// TIA Portal project "XSFW_TIA60401_A5" (V13) (continued)
   "ArrMC005" AT %T79 : Timer;   // Timer arranque MC005
   "MC004_TTB" AT %E6.3 : Bool;   // M COMPRESOR ALTA ABC4-TERMOSTATO AGUA / Compresor ABC4 Alta Temperatura de agua
   "MC005" AT %A1.2 : Bool;   // M COMPRESOR ALTA ABC5-CONTACTOR / Compresor ABC5-. Marcha-(200 Kw)
   "MC005-CO" AT %E3.5 : Bool;   // M COMPRESOR ALTA ABC5-CONFIRMACIÓN DE MARCHA / Compresor ABC5-Confirmacion Marcha-(200 Kw)
   "MC005-TO" AT %E3.6 : Bool;   // M COMPRESOR ALTA ABC5-TÉRMICO / Compresor ABC5-Falla Termico--(200 Kw)
   "MC005_EV" AT %A2.4 : Bool;   // M COMPRESOR ALTA ABC5-ELECTROVÁLVULA / Electrovalvula libera carga MC005 (ABC5)
   "MC005_MANT" AT %A3.1 : Bool;   // M COMPRESOR ALTA ABC5-SEÑAL MODO MANTENIMIENTO / Compresor MC005 Salida Mantenimiento
   "MC005_PTA" AT %E6.4 : Bool;   // M COMPRESOR ALTA ABC5-PRESOSTATO ACEITE / Compresor ABC5 Baja Presion de Aceite
   "MC005_PTB" AT %E6.5 : Bool;   // M COMPRESOR ALTA ABC5-PRESOSTATO AGUA / Compresor ABC5 Baja Presion de Agua
   "MC005_TTA" AT %E6.6 : Bool;   // M COMPRESOR ALTA ABC5-TERMOSTATO AIRE / Compresor ABC5 Alta Temperatura de Aire
   "MC005_TTB" AT %E6.7 : Bool;   // M COMPRESOR ALTA ABC5-TERMOSTATO AGUA / Compresor ABC5 Alta Temperatura de agua
   "MC060-CO" AT %E10.0 : Bool;   // M COMPR BAJA SULLAIR 2-CONFIRMACIÓN DE MARCHA / Compresor Baja XXX - Conf.Marcha
   "MC060-TO" AT %E10.1 : Bool;   // M COMPR BAJA SULLAIR 2-TÉRMICO / Compresor Baja XXX - Falla de termico
   "MC060-VS1" AT %E10.2 : Bool;   // M COMPR BAJA SULLAIR 2-PULSADOR PARADA / Compresor Baja XXX - Falla de seguridades
   "MC060_MANT" AT %A5.4 : Bool;   // M COMPR BAJA SULLAIR 2-SEÑAL MODO MANTENIMIENTO / compresor XXX salida de mantenimiento
   "MC060_MARCHA" AT %A5.5 : Bool;   // M COMPR BAJA SULLAIR 2-CONTACTOR / compresor XXX salida de marcha
   "MC061-CO" AT %E11.4 : Bool;   // M COMPR BAJA SULLAIR 1-CONFIRMACIÓN DE MARCHA / Compresor Baja SULL 1 - Conf.Marcha
   "MC003_EV" AT %A2.2 : Bool;   // M COMPRESOR ALTA BELLIS-ELECTROVÁLVULA 1 / Electrovalvula libera carga MC003 (Bellis)
   "Encendido" AT %M301.1 : Bool;   // Encendido de PLC
   "MT009-TO" AT %E66.5 : Bool;   // B INT L3 Y L5-TÉRMICO / Bomba Principal Chiller Envasado - Falla de Térmico
   "MT010-CO" AT %E66.6 : Bool;   // B INT L1 Y MANOMEC-CONFIRMACIÓN DE MARCHA / Bomba Auxilliar Chiller Envasado - Confirmación de Marcha
   "MT010-Marcha" AT %A66.3 : Bool;   // B INT L1 Y MANOMEC-CONTACTOR / Accionamiento Bomba Intercambiador LINEA 1 Y MANOMEC
   "MT010-TO" AT %E66.7 : Bool;   // B INT L1 Y MANOMEC-TÉRMICO / Bomba Auxiliar Chiller Envasado - Falla de Térmico
   "MV030" AT %A0.2 : Bool;   // M VENTILADOR 2-CONTACTOR / VENTILADOR TORRE 1 -. marcha-
   "MV030-CO" AT %E0.4 : Bool;   // M VENTILADOR 2-CONFIRMACIÓN DE MARCHA / VENTILADOR TORRE 1 -confirmacion marcha-
   "MV030-TO" AT %E0.5 : Bool;   // M VENTILADOR 2-TÉRMICO / VENTILADOR TORRE 1 -falla termico-
   "MV030_PA" AT %E8.5 : Bool;   // M VENTILADOR 2-PULSADOR MARCHA / Ventilador 1 Torre Cavalleto Pulsador Arranque
   "MV030_PP" AT %E8.6 : Bool;   // M VENTILADOR 2-PULSADOR PARADA / Ventilador 1 Torre Cavalleto Pulsador Parada
   "MV031" AT %A0.3 : Bool;   // M VENTILADOR 1-CONTACTOR / VENTILADOR TORRE 2 -. marcha-
   "MV031-CO" AT %E0.6 : Bool;   // M VENTILADOR 1-CONFIRMACIÓN DE MARCHA / VENTILADOR TORRE 2 -confirmacion marcha-
   "MV031-TO" AT %E0.7 : Bool;   // M VENTILADOR 1-TÉRMICO / VENTILADOR TORRE 2 -falla termico-
   "MV031_PA" AT %E8.7 : Bool;   // M VENTILADOR 1-PULSADOR MARCHA / Ventilador 2 Torre Cavalleto Pulsaor Arranque
   "MV031_PP" AT %E9.0 : Bool;   // M VENTILADOR 1-PULSADOR PARADA / Ventilador 2 Torre Cavalleto Pulsaor Parada
   "iGMBooster2" AT %E9.7 : Bool;   // M BOOSTER 2-GUARDAMOTOR / Guardamotor Booster 2
   "Hab-CHILL1" AT %A69.4 : Bool;   // CHILLER 1-SEÑAL A CHILLER / Deshabilitación Chiller Soplado GRANDE
   "Hab-CHILL2" AT %A69.5 : Bool;   // CHILLER 2-SEÑAL A CHILLER / Deshabilitación Chiller Soplado CHICO
   "Hab-CHILL3" AT %A69.6 : Bool;   // CHILLER 3-SEÑAL A CHILLER / Deshabilitación Chiller Envasado GRANDE
   "Hab-CHILL4" AT %A69.7 : Bool;   // CHILLER 4-SEÑAL A CHILLER / Deshabilitación Chiller Envasado CHICO
   "ILUMINACION" AT %A0.5 : Bool;   // ILUMINACION-CONTACTOR / ILUMINACION
   "MC003_ConfPurga" AT %E1.2 : Bool;   // Bellis - Confirmación de electroválvula de purga. / Iluminacion-confirmacion marcha-
   "MC004_ConfPurga" AT %E1.3 : Bool;   // ABC4 - Confirmación de electroválvula de purga. / Iluminacion Termico
   "IndicadorChillers" AT %M310.0 : Bool;   // Indicador Aviso en chillers
   "TsinReq1" AT %T52 : Timer;   // Timeout estando en estado sin requerimiento 1
   "TsinReq2" AT %T40 : Timer;   // Timeout estando en estado sin requerimiento 2
   "TsinReq3" AT %T41 : Timer;   // Timeout estando en estado sin requerimiento 3
   "TsinReq4" AT %T42 : Timer;   // Timeout estando en estado sin requerimiento 4
   "TsinReq5" AT %T43 : Timer;   // Timeout estando en estado sin requerimiento 5
   "UNO" AT %M0.1 : Bool;
   "V001-CO" AT %E76.5 : Bool;   // VENT 1 TORR ENF CHILLERS-CONFIRMACIÓN DE MARCHA / Ventilador 1 Torres Enfriamiento - Confirmación de Marcha
   "V001-Marcha" AT %A67.6 : Bool;   // VENT 1 TORR ENF CHILLERS-CONTACTOR / Accionamiento Ventilador 1 Torres Enfriamiento
   "V001-TO" AT %E76.6 : Bool;   // VENT 1 TORR ENF CHILLERS-TÉRMICO / Ventilador 1 Torres Enfriamiento - Falla de Térmico
   "V002-CO" AT %E76.7 : Bool;   // VENT 2 TORR ENF CHILLERS-CONFIRMACIÓN DE MARCHA / Ventilador 2 Torres Enfriamiento - Confirmación de Marcha
   "V002-Marcha" AT %A67.7 : Bool;   // VENT 2 TORR ENF CHILLERS-CONTACTOR / Accionamiento Ventilador 2 Torres Enfriamiento
   "V002-TO" AT %E77.0 : Bool;   // VENT 2 TORR ENF CHILLERS-TÉRMICO / Ventilador 2 Torres Enfriamiento - Falla de Térmico
   "V003-CO" AT %E77.1 : Bool;   // VENT 3 TORR ENF CHILLERS-CONFIRMACIÓN DE MARCHA / Ventilador 3 Torres Enfriamiento - Confirmación de Marcha
   "V003-Marcha" AT %A68.0 : Bool;   // VENT 3 TORR ENF CHILLERS-CONTACTOR / Accionamiento Ventilador 3 Torres Enfriamiento
   "V003-TO" AT %E77.2 : Bool;   // VENT 3 TORR ENF CHILLERS-TÉRMICO / Ventilador 3 Torres Enfriamiento - Falla de Térmico
   "FlancoNSop1" AT %M326.1 : Bool;
   "FlancoNSop2" AT %M326.2 : Bool;
   "FlancoNSop3" AT %M326.3 : Bool;
   "FlancoNoFaGen" AT %M325.2 : Bool;
   "FlancoNoFal1" AT %M324.5 : Bool;
   "MC003_EV2" AT %A3.2 : Bool;   // M COMPRESOR ALTA BELLIS-ELECTROVÁLVULA 2 / Electrovalvula media carga Bellis
   "MC003_FTA" AT %E7.4 : Bool;   // M COMPRESOR ALTA BELLIS-FUJOSTATO / Compresor Bellis & MHW28 Falla de Flujostato
   "MC003_MANT" AT %A2.7 : Bool;   // M COMPRESOR ALTA BELLIS-SEÑAL MODO MANTENIMIENTO / Compresor MC003 Salida Mantenimiento
   "MC003_PTA" AT %E7.0 : Bool;   // M COMPRESOR ALTA BELLIS-PRESOSTATO ACEITE / Compresor Bellis & MHW28 Baja Presion Aceite
   "MC003_PTB" AT %E7.1 : Bool;   // M COMPRESOR ALTA BELLIS-PRESOSTATO AGUA / Compresor Bellis & MHW28 Baja Presion de Agua
   "MC003_TTA" AT %E7.2 : Bool;   // M COMPRESOR ALTA BELLIS-TERMOSTATO AIRE / Compresor Bellis & MHW28 Alta temperatura de Aire
   "MC003_TTB" AT %E7.3 : Bool;   // M COMPRESOR ALTA BELLIS-TERMOSTATO AGUA / Compresor Bellis & MHW28 Alta temperatura de Agua
   "MC004" AT %A1.1 : Bool;   // M COMPRESOR ALTA ABC4-CONTACTOR / Compresor ABC4-. Marcha-
   "MC004-CO" AT %E3.3 : Bool;   // M COMPRESOR ALTA ABC4-CONFIRMACIÓN DE MARCHA / Compresor ABC4-Confirmacion Marcha-
   "MC004-TO" AT %E3.4 : Bool;   // M COMPRESOR ALTA ABC4-TÉRMICO / Compresor ABC4-Falla Termico-
   "MC004_EV" AT %A2.3 : Bool;   // M COMPRESOR ALTA ABC4-ELECTROVÁLVULA / Electrovalvula libera carga MC004 (ABC4)
   "MC004_MANT" AT %A3.0 : Bool;   // M COMPRESOR ALTA ABC4-SEÑAL MODO MANTENIMIENTO / Compresor MC004 Salida Mantenimiento
   "MC004_PTA" AT %E6.0 : Bool;   // M COMPRESOR ALTA ABC4-PRESOSTATO ACEITE / Compresor ABC4 Baja Presion de Aceite
   "MC004_PTB" AT %E6.1 : Bool;   // M COMPRESOR ALTA ABC4-PRESOSTATO AGUA / Compresor ABC4 Baja Presion de Agua
   "MC004_TTA" AT %E6.2 : Bool;   // M COMPRESOR ALTA ABC4-TERMOSTATO AIRE / Compresor ABC4 Alta Temperatura de Aire
   "MC001_PTA" AT %E5.0 : Bool;   // M COMPRESOR ALTA ABC2-PRESOSTATO ACEITE / Compresor ABC2 Baja Presion de Aceite
   "MC001_PTB" AT %E5.1 : Bool;   // M COMPRESOR ALTA ABC2-PRESOSTATO AGUA / Compresor ABC2 Baja Presion de Agua
   "MC001_TTA" AT %E5.2 : Bool;   // M COMPRESOR ALTA ABC2-TERMOSTATO AIRE / Compresor ABC2 Alta Temperatura de Aire
   "MC001_TTB" AT %E5.3 : Bool;   // M COMPRESOR ALTA ABC2-TERMOSTATO AGUA / Compresor ABC2 Alta Temperatura de agua
   "MC002" AT %A0.7 : Bool;   // M COMPRESOR ALTA ABC3-CONTACTOR / Compresor ABC3-. Marcha-
   "MC002-CO" AT %E2.7 : Bool;   // M COMPRESOR ALTA ABC3-CONFIRMACIÓN DE MARCHA / Compresor ABC3-Confirmacion Marcha-
   "MC002-TO" AT %E3.0 : Bool;   // M COMPRESOR ALTA ABC3-TÉRMICO / Compresor ABC3-Falla Termico-
   "MC002_EV" AT %A2.1 : Bool;   // M COMPRESOR ALTA ABC3-ELECTROVÁLVULA / Electrovalvula libera carga MC002 (ABC3)
   "MC002_MANT" AT %A2.6 : Bool;   // M COMPRESOR ALTA ABC3-SEÑAL MODO MANTENIMIENTO / Compresor MC002 Salida Mantenimiento
   "MC002_PTA" AT %E5.4 : Bool;   // M COMPRESOR ALTA ABC3-PRESOSTATO ACEITE / Compresor ABC3 Baja Presion de Aceite
   "MC002_PTB" AT %E5.5 : Bool;   // M COMPRESOR ALTA ABC3-PRESOSTATO AGUA / Compresor ABC3 Baja Presion de Agua
   "MC002_TTA" AT %E5.6 : Bool;   // M COMPRESOR ALTA ABC3-TERMOSTATO AIRE / Compresor ABC3 Alta Temperatura de Aire
   "MC002_TTB" AT %E5.7 : Bool;   // M COMPRESOR ALTA ABC3-TERMOSTATO AGUA / Compresor ABC3 Alta Temperatura de agua
   "MC003" AT %A1.0 : Bool;   // M COMPRESOR ALTA BELLIS-CONTACTOR / Compresor B&MWH28-. Marcha-
   "MC003-CO" AT %E3.1 : Bool;   // M COMPRESOR ALTA BELLIS-CONFIRMACIÓN DE MARCHA / Compresor B&MWH28-Confirmacion Marcha-
   "MC003-TO" AT %E3.2 : Bool;   // M COMPRESOR ALTA BELLIS-TÉRMICO / Compresor B&MWH28-Falla Termico-
   "BoostPlsManual" AT %M10.6 : Bool;   // Booster Pulsa Manual desde HMI
   "BoostPlsAutoma" AT %M10.7 : Bool;   // Booster Pulsa Automático desde HMI
   "ErrPMQG" AT %M321.2 : Bool;   // Error Prioritarias General
   "PRESOSTATO-TORRES" AT %E76.4 : Bool;   // CHILLER (TODOS)-PRESOSTATO / Presostato Agua Torres de Enfriamiento
   "PT2_AIRE" AT %E4.7 : Bool;   // - / PRESOSTATO ALTA PRESION DE AIRE EN COLECTOR 40Kg
   "Parada-MC061" AT %A6.1 : Bool;   // M COMPR BAJA SULLAIR 1-ORDEN PARADA / Parada MC061
   "MC006_ConfPurga" AT %E11.7 : Bool;   // ABC1 - Confirmación de electroválvula de purga.
   "MP014-TO" AT %E0.1 : Bool;   // BOMBA 1-TÉRMICO / BOMBA 1TORRE ENF.-TERMICO
   "MP015" AT %A0.1 : Bool;   // BOMBA 2-CONTACTOR / BOMBA 2 TORRE -. marcha-
   "MP015-CO" AT %E0.2 : Bool;   // BOMBA 2-CONFIRMACIÓN DE MARCHA / BOMBA 2 TORRE ENF.-CONFIRMACION
   "MP015-TO" AT %E0.3 : Bool;   // BOMBA 2-TÉRMICO / BOMBA 2 TORRE ENF.-TERMICO
   "MP018-CO" AT %E68.0 : Bool;   // BOMBA 1-CONFIRMACIÓN DE MARCHA / Bomba 1 Torres Enfriamiento - Confirmación de Marcha
   "MP018-Marcha" AT %A67.0 : Bool;   // BOMBA 1-CONTACTOR / Accionamiento Bomba 1 Torres Enfriamiento
   "MP018-TO" AT %E68.1 : Bool;   // BOMBA 1-TÉRMICO / Bomba 1 Torres Enfriamiento - Falla de Térmico
   "MP018_PA" AT %E8.1 : Bool;   // BOMBA 1-PULSADOR MARCHA / Bomba 1 Torre Cavalleto Pulsador Arranque
   "MP018_PP" AT %E8.2 : Bool;   // BOMBA 1-PULSADOR PARADA / Bomba 1 Torre Cavalleto Pulsador Parada
   "MC001_ConfPurga" AT %E1.0 : Bool;   // ABC2 - Confirmación de electroválvula de purga. / Bomba de pozo -confirmacion marcha-
   "CERO" AT %M0.0 : Bool;
   "CHILL1-AL1" AT %E68.4 : Bool;   // CHILLER SOPLADO-ALARMA 1 / Chiller Soplado GRANDE - Alarma 1
   "CHILL1-AL2" AT %E68.5 : Bool;   // CHILLER SOPLADO-ALARMA 2 / Chiller Soplado GRANDE - Alarma 2
   "CHILL1-MAX" AT %E68.7 : Bool;   // CHILLER SOPLADO-MAXIMA CAPACIDAD / Chiller Soplado GRANDE - Máxima Capacidad
   "CHILL1-RUN" AT %E68.6 : Bool;   // CHILLER SOPLADO- / Chiller Soplado GRANDE - En modo RUN
   "CHILL2-" AT %E69.0 : Bool;   // CHILLER SOPLADO CHICO- / Chiller Soplado CHICO - Contactor 1
   "CHILL2-b" AT %E69.1 : Bool;   // CHILLER SOPLADO CHICO- / Chiller Soplado CHICO - Contactor 2
   "CHILL2-c" AT %E69.2 : Bool;   // CHILLER SOPLADO CHICO-FALLA / Chiller Soplado CHICO - Termico Contactor 1
   "CHILL2-d" AT %E69.3 : Bool;   // CHILLER SOPLADO CHICO-FALLA / Chiller Soplado CHICO - Termico Contactor 2
   "CHILL3-AL1" AT %E69.4 : Bool;   // CHILLER ENVASADO GRAND-ALARMA 1 / Chiller Envasado GRANDE - Alarma 1
   "MC064-VS1" AT %E11.3 : Bool;   // M COMPR BAJA ATLAS 2-PULSADOR PARADA / Compresor Baja ATLAS 2 - Falla de seguridades
   "MC064_MANT" AT %A5.2 : Bool;   // M COMPR BAJA ATLAS 2-SEÑAL MODO MANTENIMIENTO / compresor ATLAS 2 salida de mantenimiento
   "MC064_MARCHA" AT %A5.3 : Bool;   // M COMPR BAJA ATLAS 2-CONTACTOR / compresor ATLAS 2 salida de marcha
   "MP010-CO" AT %E67.0 : Bool;   // B PRINC CH. SOPLADO-CONFIRMACIÓN DE MARCHA / Bomba Intercambiador LINEA 1 - Confirmación de Marcha
   "MP010-Marcha" AT %A66.4 : Bool;   // B PRINC CH. SOPLADO-CONTACTOR / Accionamiento Bomba Principal Chiller Soplado
   "MP010-TO" AT %E67.1 : Bool;   // B PRINC CH. SOPLADO-TÉRMICO / Bomba Intercambiador LINEA 1 - Falla de Térmico
   "MC006" AT %Q6.2 : Bool;   // M COMPRESOR ALTA ABC1-CONTACTOR
   "MC006_EV" AT %Q6.3 : Bool;   // M COMPRESOR ALTA ABC1-ELECTROVÁLVULA
   "MC006_MANT" AT %Q6.4 : Bool;   // M COMPRESOR ALTA ABC1-SEÑAL MODO MANTENIMIENTO
   "TsinReq6" AT %T59 : Timer;
   "TV6" AT %T69 : Timer;
   "flReqMch6" AT %M0.5 : Bool;
   "ErrPMQ6" AT %M1.5 : Bool;
   "ErrCMQ6" AT %M1.6 : Bool;
   "RetVLV6" AT %T85 : Timer;
   "TRetVCmp6" AT %T86 : Timer;
   "ArrMC006" AT %T88 : Timer;
   "FlaAux6" AT %M301.2 : Bool;
   "FlancoINC6" AT %M326.7 : Bool;
   "FlancoDEC6" AT %M327.0 : Bool;
   "FlancoMan6" AT %M327.1 : Bool;
   "FlancoManP6" AT %M327.2 : Bool;
   "FlancoAuto6" AT %M327.3 : Bool;
   "FlancoNoFal6" AT %M327.4 : Bool;
   "FlancoTSinReq6" AT %M327.5 : Bool;
   "AuxTempMS050" AT %MW340 : Int;
   "AuxTempMS051" AT %MW342 : Int;
   "AuxTempMS052" AT %MW344 : Int;
   "AuxTempMS053" AT %MW346 : Int;
   "AuxTempMS054" AT %MW348 : Int;
   "AuxTempMS055" AT %MW350 : Int;
   "AuxTempMS056" AT %MW352 : Int;
   "AuxTempMC060" AT %MW354 : Int;
   "AuxTempMC061" AT %MW356 : Int;
   "AuxTempMC062" AT %MW358 : Int;
   "AuxTempMC063" AT %MW360 : Int;
   "AuxTempMC064" AT %MW362 : Int;
   "AuxTempMC065" AT %MW364 : Int;
   "ProxMantBoost1" AT %MD16 : DInt;
   "LimiteMantBoost1" AT %M1.7 : Bool;
   "ProxMantBoost2" AT %MD26 : DInt;
   "LimiteMantBoost2" AT %M2.3 : Bool;
END_VAR

DATA_BLOCK "DB_Fecha"   // DB1
{ S7_Optimized_Access := 'FALSE' }
VERSION : 0.1
   VAR
      STAT0 : Date_And_Time;
      STAT1 : Int;
      STAT2 : Int;
      STAT3 : Int;
      STAT4 : Int;
      STAT5 : Int;
      STAT6 : Int;
      STAT7 : Int;
      STAT8 : Int;
      STAT9 : Int;
      STAT10 : Int;
      STAT11 : Word;
      STAT12 : Word;
      STAT13 : Word;
      STAT14 : Word;
      STAT15 : Word;
      STAT16 : Word;
   END_VAR
BEGIN
END_DATA_BLOCK

DATA_BLOCK "Enclavamientos"   // DB28
{ S7_Optimized_Access := 'FALSE' }
VERSION : 0.1
   VAR
      En1 : Bool;
      En2 : Bool;
      En3 : Bool;
      En4 : Bool;
      En5 : Bool;
      En6 : Bool;
      En7 : Bool;
      En8 : Bool;
      En9 : Bool;
      En10 : Bool;
      En11 : Bool;
      En12 : Bool;
      En13 : Bool;
      En14 : Bool;
      En15 : Bool;
      En16 : Bool;
      En17 : Bool;
      En18 : Bool;
      En19 : Bool;
      En20 : Bool;
      En21 : Bool;
      En22 : Bool;
      En23 : Bool;
      En24 : Bool;
      En25 : Bool;
      En26 : Bool;
      En27 : Bool;
      En28 : Bool;
      En29 : Bool;
      En30 : Bool;
      En31 : Bool;
      En32 : Bool;
      En33 : Bool;
      En34 : Bool;
      En35 : Bool;
      En36 : Bool;
      En37 : Bool;
      En38 : Bool;
      En39 : Bool;
      En40 : Bool;
      En41 : Bool;
      En42 : Bool;
      En43 : Bool;
      En44 : Bool;
      En45 : Bool;
      En46 : Bool;
      En47 : Bool;
      En48 : Bool;
      En49 : Bool;
      En50 : Bool;
      En51 : Bool;
      En52 : Bool;
      En53 : Bool;
      En54 : Bool;
      En55 : Bool;
      En56 : Bool;
      En57 : Bool;
      En58 : Bool;
      En59 : Bool;
      En60 : Bool;
      En61 : Bool;
      En62 : Bool;
      En63 : Bool;
      En64 : Bool;
   END_VAR
BEGIN
END_DATA_BLOCK

// folder: Alarmas

DATA_BLOCK "DB_ALA_PRE"   // DB32
{ S7_Optimized_Access := 'FALSE' }
VERSION : 0.1
   VAR
      x : Bool;
      x1 : Bool;
      x2 : Bool;
      x3 : Bool;
      x4 : Bool;
      x5 : Bool;
      x6 : Bool;
      x7 : Bool;
      x8 : Bool;
      x9 : Bool;
      x10 : Bool;
      x11 : Bool;
      x12 : Bool;
      x13 : Bool;
      x14 : Bool;
      x15 : Bool;
      x16 : Bool;
      x17 : Bool;
      x18 : Bool;
      x19 : Bool;
      x20 : Bool;
      x21 : Bool;
      x22 : Bool;
      x23 : Bool;
      x24 : Bool;
      x25 : Bool;
      x26 : Bool;
      x27 : Bool;
      x28 : Bool;
      x29 : Bool;
      x30 : Bool;
      x31 : Bool;
      x32 : Bool;
      x33 : Bool;
      x34 : Bool;
      x35 : Bool;
      x36 : Bool;
      x37 : Bool;
      x38 : Bool;
      x39 : Bool;
      x40 : Bool;
      x41 : Bool;
      x42 : Bool;
      x43 : Bool;
      x44 : Bool;
      x45 : Bool;
      x46 : Bool;
      x47 : Bool;
      x48 : Bool;
      x49 : Bool;
      x50 : Bool;
      x51 : Bool;
      x52 : Bool;
      x53 : Bool;
      x54 : Bool;
      x55 : Bool;
      x56 : Bool;
      x57 : Bool;
      x58 : Bool;
      x59 : Bool;
      x60 : Bool;
      x61 : Bool;
      x62 : Bool;
      x63 : Bool;
      x64 : Bool;
      x65 : Bool;
      x66 : Bool;
      x67 : Bool;
      x68 : Bool;
      x69 : Bool;
      x70 : Bool;
      x71 : Bool;
      x72 : Bool;
      x73 : Bool;
      x74 : Bool;
      x75 : Bool;
      x76 : Bool;
      x77 : Bool;
      x78 : Bool;
      x79 : Bool;
      x80 : Bool;
      x81 : Bool;
      x82 : Bool;
      x83 : Bool;
      x84 : Bool;
      x85 : Bool;
      x86 : Bool;
      x87 : Bool;
      x88 : Bool;
      x89 : Bool;
      x90 : Bool;
      x91 : Bool;
      x92 : Bool;
      x93 : Bool;
      x94 : Bool;
      x95 : Bool;
      x96 : Bool;
      x97 : Bool;
      x98 : Bool;
      x99 : Bool;
      x100 : Bool;
      x101 : Bool;
      x102 : Bool;
      x103 : Bool;
      x104 : Bool;
      x105 : Bool;
      x106 : Bool;
      x107 : Bool;
      x108 : Bool;
      x109 : Bool;
      x110 : Bool;
      x111 : Bool;
      x112 : Bool;
      x113 : Bool;
      x114 : Bool;
      x115 : Bool;
      x116 : Bool;
      x117 : Bool;
      x118 : Bool;
      x119 : Bool;
      x120 : Bool;
      x121 : Bool;
      x122 : Bool;
      x123 : Bool;
      x124 : Bool;
      x125 : Bool;
      x126 : Bool;
      x127 : Bool;
      x128 : Bool;
      x129 : Bool;
      x130 : Bool;
      x131 : Bool;
      x132 : Bool;
      x133 : Bool;
      x134 : Bool;
      x135 : Bool;
      x136 : Bool;
      x137 : Bool;
      x138 : Bool;
      x139 : Bool;
      x140 : Bool;
      x141 : Bool;
      x142 : Bool;
      x143 : Bool;
      x144 : Bool;
      x145 : Bool;
      x146 : Bool;
      x147 : Bool;
      x148 : Bool;
      x149 : Bool;
      x150 : Bool;
      x151 : Bool;
      x152 : Bool;
      x153 : Bool;
      x154 : Bool;
      x155 : Bool;
      x156 : Bool;
      x157 : Bool;
      x158 : Bool;
      x159 : Bool;
      x160 : Bool;
      x161 : Bool;
      x162 : Bool;
      x163 : Bool;
      x164 : Bool;
      x165 : Bool;
      x166 : Bool;
      x167 : Bool;
      x168 : Bool;
      x169 : Bool;
      x170 : Bool;
      x171 : Bool;
      x172 : Bool;
      x173 : Bool;
      x174 : Bool;
      x175 : Bool;
      x176 : Bool;
      x177 : Bool;
      x178 : Bool;
      x179 : Bool;
      x180 : Bool;
      x181 : Bool;
      x182 : Bool;
      x183 : Bool;
      x184 : Bool;
      x185 : Bool;
      x186 : Bool;
      x187 : Bool;
      x188 : Bool;
      x189 : Bool;
      x190 : Bool;
      x191 : Bool;
      x192 : Bool;
      x193 : Bool;
      x194 : Bool;
      x195 : Bool;
      x196 : Bool;
      x197 : Bool;
      x198 : Bool;
      x199 : Bool;
   END_VAR
BEGIN
END_DATA_BLOCK

DATA_BLOCK "DB_ALA_REC"   // DB33
{ S7_Optimized_Access := 'FALSE' }
VERSION : 0.1
   VAR
      x : Bool;
      x1 : Bool;
      x2 : Bool;
      x3 : Bool;
      x4 : Bool;
      x5 : Bool;
      x6 : Bool;
      x7 : Bool;
      x8 : Bool;
      x9 : Bool;
      x10 : Bool;
      x11 : Bool;
      x12 : Bool;
      x13 : Bool;
      x14 : Bool;
      x15 : Bool;
      x16 : Bool;
      x17 : Bool;
      x18 : Bool;
      x19 : Bool;
      x20 : Bool;
      x21 : Bool;
      x22 : Bool;
      x23 : Bool;
      x24 : Bool;
      x25 : Bool;
      x26 : Bool;
      x27 : Bool;
      x28 : Bool;
      x29 : Bool;
      x30 : Bool;
      x31 : Bool;
      x32 : Bool;
      x33 : Bool;
      x34 : Bool;
      x35 : Bool;
      x36 : Bool;
      x37 : Bool;
      x38 : Bool;
      x39 : Bool;
      x40 : Bool;
      x41 : Bool;
      x42 : Bool;
      x43 : Bool;
      x44 : Bool;
      x45 : Bool;
      x46 : Bool;
      x47 : Bool;
      x48 : Bool;
      x49 : Bool;
      x50 : Bool;
      x51 : Bool;
      x52 : Bool;
      x53 : Bool;
      x54 : Bool;
      x55 : Bool;
      x56 : Bool;
      x57 : Bool;
      x58 : Bool;
      x59 : Bool;
      x60 : Bool;
      x61 : Bool;
      x62 : Bool;
      x63 : Bool;
      x64 : Bool;
      x65 : Bool;
      x66 : Bool;
      x67 : Bool;
      x68 : Bool;
      x69 : Bool;
      x70 : Bool;
      x71 : Bool;
      x72 : Bool;
      x73 : Bool;
      x74 : Bool;
      x75 : Bool;
      x76 : Bool;
      x77 : Bool;
      x78 : Bool;
      x79 : Bool;
      x80 : Bool;
      x81 : Bool;
      x82 : Bool;
      x83 : Bool;
      x84 : Bool;
      x85 : Bool;
      x86 : Bool;
      x87 : Bool;
      x88 : Bool;
      x89 : Bool;
      x90 : Bool;
      x91 : Bool;
      x92 : Bool;
      x93 : Bool;
      x94 : Bool;
      x95 : Bool;
      x96 : Bool;
      x97 : Bool;
      x98 : Bool;
      x99 : Bool;
      x100 : Bool;
      x101 : Bool;
      x102 : Bool;
      x103 : Bool;
      x104 : Bool;
      x105 : Bool;
      x106 : Bool;
      x107 : Bool;
      x108 : Bool;
      x109 : Bool;
      x110 : Bool;
      x111 : Bool;
      x112 : Bool;
      x113 : Bool;
      x114 : Bool;
      x115 : Bool;
      x116 : Bool;
      x117 : Bool;
      x118 : Bool;
      x119 : Bool;
      x120 : Bool;
      x121 : Bool;
      x122 : Bool;
      x123 : Bool;
      x124 : Bool;
      x125 : Bool;
      x126 : Bool;
      x127 : Bool;
      x128 : Bool;
      x129 : Bool;
      x130 : Bool;
      x131 : Bool;
      x132 : Bool;
      x133 : Bool;
      x134 : Bool;
      x135 : Bool;
      x136 : Bool;
      x137 : Bool;
      x138 : Bool;
      x139 : Bool;
      x140 : Bool;
      x141 : Bool;
      x142 : Bool;
      x143 : Bool;
      x144 : Bool;
      x145 : Bool;
      x146 : Bool;
      x147 : Bool;
      x148 : Bool;
      x149 : Bool;
      x150 : Bool;
      x151 : Bool;
      x152 : Bool;
      x153 : Bool;
      x154 : Bool;
      x155 : Bool;
      x156 : Bool;
      x157 : Bool;
      x158 : Bool;
      x159 : Bool;
      x160 : Bool;
      x161 : Bool;
      x162 : Bool;
      x163 : Bool;
      x164 : Bool;
      x165 : Bool;
      x166 : Bool;
      x167 : Bool;
      x168 : Bool;
      x169 : Bool;
      x170 : Bool;
      x171 : Bool;
      x172 : Bool;
      x173 : Bool;
      x174 : Bool;
      x175 : Bool;
      x176 : Bool;
      x177 : Bool;
      x178 : Bool;
      x179 : Bool;
      x180 : Bool;
      x181 : Bool;
      x182 : Bool;
      x183 : Bool;
      x184 : Bool;
      x185 : Bool;
      x186 : Bool;
      x187 : Bool;
      x188 : Bool;
      x189 : Bool;
      x190 : Bool;
      x191 : Bool;
      x192 : Bool;
      x193 : Bool;
      x194 : Bool;
      x195 : Bool;
      x196 : Bool;
      x197 : Bool;
      x198 : Bool;
      x199 : Bool;
   END_VAR
BEGIN
END_DATA_BLOCK

DATA_BLOCK "DB_ALA_MEM"   // DB34
{ S7_Optimized_Access := 'FALSE' }
VERSION : 0.1
   VAR
      x : Bool;
      x1 : Bool;
      x2 : Bool;
      x3 : Bool;
      x4 : Bool;
      x5 : Bool;
      x6 : Bool;
      x7 : Bool;
      x8 : Bool;
      x9 : Bool;
      x10 : Bool;
      x11 : Bool;
      x12 : Bool;
      x13 : Bool;
      x14 : Bool;
      x15 : Bool;
      x16 : Bool;
      x17 : Bool;
      x18 : Bool;
      x19 : Bool;
      x20 : Bool;
      x21 : Bool;
      x22 : Bool;
      x23 : Bool;
      x24 : Bool;
      x25 : Bool;
      x26 : Bool;
      x27 : Bool;
      x28 : Bool;
      x29 : Bool;
      x30 : Bool;
      x31 : Bool;
      x32 : Bool;
      x33 : Bool;
      x34 : Bool;
      x35 : Bool;
      x36 : Bool;
      x37 : Bool;
      x38 : Bool;
      x39 : Bool;
      x40 : Bool;
      x41 : Bool;
      x42 : Bool;
      x43 : Bool;
      x44 : Bool;
      x45 : Bool;
      x46 : Bool;
      x47 : Bool;
      x48 : Bool;
      x49 : Bool;
      x50 : Bool;
      x51 : Bool;
      x52 : Bool;
      x53 : Bool;
      x54 : Bool;
      x55 : Bool;
      x56 : Bool;
      x57 : Bool;
      x58 : Bool;
      x59 : Bool;
      x60 : Bool;
      x61 : Bool;
      x62 : Bool;
      x63 : Bool;
      x64 : Bool;
      x65 : Bool;
      x66 : Bool;
      x67 : Bool;
      x68 : Bool;
      x69 : Bool;
      x70 : Bool;
      x71 : Bool;
      x72 : Bool;
      x73 : Bool;
      x74 : Bool;
      x75 : Bool;
      x76 : Bool;
      x77 : Bool;
      x78 : Bool;
      x79 : Bool;
      x80 : Bool;
      x81 : Bool;
      x82 : Bool;
      x83 : Bool;
      x84 : Bool;
      x85 : Bool;
      x86 : Bool;
      x87 : Bool;
      x88 : Bool;
      x89 : Bool;
      x90 : Bool;
      x91 : Bool;
      x92 : Bool;
      x93 : Bool;
      x94 : Bool;
      x95 : Bool;
      x96 : Bool;
      x97 : Bool;
      x98 : Bool;
      x99 : Bool;
      x100 : Bool;
      x101 : Bool;
      x102 : Bool;
      x103 : Bool;
      x104 : Bool;
      x105 : Bool;
      x106 : Bool;
      x107 : Bool;
      x108 : Bool;
      x109 : Bool;
      x110 : Bool;
      x111 : Bool;
      x112 : Bool;
      x113 : Bool;
      x114 : Bool;
      x115 : Bool;
      x116 : Bool;
      x117 : Bool;
      x118 : Bool;
      x119 : Bool;
      x120 : Bool;
      x121 : Bool;
      x122 : Bool;
      x123 : Bool;
      x124 : Bool;
      x125 : Bool;
      x126 : Bool;
      x127 : Bool;
      x128 : Bool;
      x129 : Bool;
      x130 : Bool;
      x131 : Bool;
      x132 : Bool;
      x133 : Bool;
      x134 : Bool;
      x135 : Bool;
      x136 : Bool;
      x137 : Bool;
      x138 : Bool;
      x139 : Bool;
      x140 : Bool;
      x141 : Bool;
      x142 : Bool;
      x143 : Bool;
      x144 : Bool;
      x145 : Bool;
      x146 : Bool;
      x147 : Bool;
      x148 : Bool;
      x149 : Bool;
      x150 : Bool;
      x151 : Bool;
      x152 : Bool;
      x153 : Bool;
      x154 : Bool;
      x155 : Bool;
      x156 : Bool;
      x157 : Bool;
      x158 : Bool;
      x159 : Bool;
      x160 : Bool;
      x161 : Bool;
      x162 : Bool;
      x163 : Bool;
      x164 : Bool;
      x165 : Bool;
      x166 : Bool;
      x167 : Bool;
      x168 : Bool;
      x169 : Bool;
      x170 : Bool;
      x171 : Bool;
      x172 : Bool;
      x173 : Bool;
      x174 : Bool;
      x175 : Bool;
      x176 : Bool;
      x177 : Bool;
      x178 : Bool;
      x179 : Bool;
      x180 : Bool;
      x181 : Bool;
      x182 : Bool;
      x183 : Bool;
      x184 : Bool;
      x185 : Bool;
      x186 : Bool;
      x187 : Bool;
      x188 : Bool;
      x189 : Bool;
      x190 : Bool;
      x191 : Bool;
      x192 : Bool;
      x193 : Bool;
      x194 : Bool;
      x195 : Bool;
      x196 : Bool;
      x197 : Bool;
      x198 : Bool;
      x199 : Bool;
   END_VAR
BEGIN
END_DATA_BLOCK

DATA_BLOCK "DB_COM_REC"   // DB35
{ S7_Optimized_Access := 'FALSE' }
VERSION : 0.1
   VAR
      x : Bool;
      x1 : Bool;
      x2 : Bool;
      x3 : Bool;
      x4 : Bool;
      x5 : Bool;
      x6 : Bool;
      x7 : Bool;
      x8 : Bool;
      x9 : Bool;
      x10 : Bool;
      x11 : Bool;
      x12 : Bool;
      x13 : Bool;
      x14 : Bool;
      x15 : Bool;
      x16 : Bool;
      x17 : Bool;
      x18 : Bool;
      x19 : Bool;
      x20 : Bool;
      x21 : Bool;
      x22 : Bool;
      x23 : Bool;
      x24 : Bool;
      x25 : Bool;
      x26 : Bool;
      x27 : Bool;
      x28 : Bool;
      x29 : Bool;
      x30 : Bool;
      x31 : Bool;
      x32 : Bool;
      x33 : Bool;
      x34 : Bool;
      x35 : Bool;
      x36 : Bool;
      x37 : Bool;
      x38 : Bool;
      x39 : Bool;
      x40 : Bool;
      x41 : Bool;
      x42 : Bool;
      x43 : Bool;
      x44 : Bool;
      x45 : Bool;
      x46 : Bool;
      x47 : Bool;
      x48 : Bool;
      x49 : Bool;
      x50 : Bool;
      x51 : Bool;
      x52 : Bool;
      x53 : Bool;
      x54 : Bool;
      x55 : Bool;
      x56 : Bool;
      x57 : Bool;
      x58 : Bool;
      x59 : Bool;
      x60 : Bool;
      x61 : Bool;
      x62 : Bool;
      x63 : Bool;
      x64 : Bool;
      x65 : Bool;
      x66 : Bool;
      x67 : Bool;
      x68 : Bool;
      x69 : Bool;
      x70 : Bool;
      x71 : Bool;
      x72 : Bool;
      x73 : Bool;
      x74 : Bool;
      x75 : Bool;
      x76 : Bool;
      x77 : Bool;
      x78 : Bool;
      x79 : Bool;
      x80 : Bool;
      x81 : Bool;
      x82 : Bool;
      x83 : Bool;
      x84 : Bool;
      x85 : Bool;
      x86 : Bool;
      x87 : Bool;
      x88 : Bool;
      x89 : Bool;
      x90 : Bool;
      x91 : Bool;
      x92 : Bool;
      x93 : Bool;
      x94 : Bool;
      x95 : Bool;
      x96 : Bool;
      x97 : Bool;
      x98 : Bool;
      x99 : Bool;
      x100 : Bool;
      x101 : Bool;
      x102 : Bool;
      x103 : Bool;
      x104 : Bool;
      x105 : Bool;
      x106 : Bool;
      x107 : Bool;
      x108 : Bool;
      x109 : Bool;
      x110 : Bool;
      x111 : Bool;
      x112 : Bool;
      x113 : Bool;
      x114 : Bool;
      x115 : Bool;
      x116 : Bool;
      x117 : Bool;
      x118 : Bool;
      x119 : Bool;
      x120 : Bool;
      x121 : Bool;
      x122 : Bool;
      x123 : Bool;
      x124 : Bool;
      x125 : Bool;
      x126 : Bool;
      x127 : Bool;
      x128 : Bool;
      x129 : Bool;
      x130 : Bool;
      x131 : Bool;
      x132 : Bool;
      x133 : Bool;
      x134 : Bool;
      x135 : Bool;
      x136 : Bool;
      x137 : Bool;
      x138 : Bool;
      x139 : Bool;
      x140 : Bool;
      x141 : Bool;
      x142 : Bool;
      x143 : Bool;
      x144 : Bool;
      x145 : Bool;
      x146 : Bool;
      x147 : Bool;
      x148 : Bool;
      x149 : Bool;
      x150 : Bool;
      x151 : Bool;
      x152 : Bool;
      x153 : Bool;
      x154 : Bool;
      x155 : Bool;
      x156 : Bool;
      x157 : Bool;
      x158 : Bool;
      x159 : Bool;
      x160 : Bool;
      x161 : Bool;
      x162 : Bool;
      x163 : Bool;
      x164 : Bool;
      x165 : Bool;
      x166 : Bool;
      x167 : Bool;
      x168 : Bool;
      x169 : Bool;
      x170 : Bool;
      x171 : Bool;
      x172 : Bool;
      x173 : Bool;
      x174 : Bool;
      x175 : Bool;
      x176 : Bool;
      x177 : Bool;
      x178 : Bool;
      x179 : Bool;
      x180 : Bool;
      x181 : Bool;
      x182 : Bool;
      x183 : Bool;
      x184 : Bool;
      x185 : Bool;
      x186 : Bool;
      x187 : Bool;
      x188 : Bool;
      x189 : Bool;
      x190 : Bool;
      x191 : Bool;
      x192 : Bool;
      x193 : Bool;
      x194 : Bool;
      x195 : Bool;
      x196 : Bool;
      x197 : Bool;
      x198 : Bool;
      x199 : Bool;
   END_VAR
BEGIN
END_DATA_BLOCK

DATA_BLOCK "DB_COM__REC_FLANCO"   // DB36
{ S7_Optimized_Access := 'FALSE' }